
       //H1
       "DB_M256F_Scada".tAlm.tS.tS0.x0 := "M256_Manag_IDB".M256F_IDB[0].tALM.tS.x0;
       "DB_M256F_Scada".tAlm.tS.tS0.x1 := "M256_Manag_IDB".M256F_IDB[0].tALM.tS.x1;
       "DB_M256F_Scada".tAlm.tS.tS0.x2 := "M256_Manag_IDB".M256F_IDB[0].tALM.tS.x2;
       "DB_M256F_Scada".tAlm.tS.tS0.x3 := "M256_Manag_IDB".M256F_IDB[0].tALM.tS.x3;
       "DB_M256F_Scada".tAlm.tS.tS0.x4 := "M256_Manag_IDB".M256F_IDB[0].tALM.tS.x4;
       "DB_M256F_Scada".tAlm.tS.tS0.x5 := "M256_Manag_IDB".M256F_IDB[0].tALM.tS.x5;
       "DB_M256F_Scada".tAlm.tS.tS0.x6 := "M256_Manag_IDB".M256F_IDB[0].tALM.tS.x6;
       "DB_M256F_Scada".tAlm.tS.tS0.x7 := "M256_Manag_IDB".M256F_IDB[0].tALM.tS.x7;
       "DB_M256F_Scada".tAlm.tS.tS0.x8 := "M256_Manag_IDB".M256F_IDB[0].tALM.tS.x8;
       //H2
       "DB_M256F_Scada".tAlm.tS.tS0.x9 := "M256_Manag_IDB".M256F_IDB[1].tALM.tS.x0;
       "DB_M256F_Scada".tAlm.tS.tS0.x10 := "M256_Manag_IDB".M256F_IDB[1].tALM.tS.x1;
       "DB_M256F_Scada".tAlm.tS.tS0.x11 := "M256_Manag_IDB".M256F_IDB[1].tALM.tS.x2;
       "DB_M256F_Scada".tAlm.tS.tS0.x12 := "M256_Manag_IDB".M256F_IDB[1].tALM.tS.x3;
       "DB_M256F_Scada".tAlm.tS.tS0.x13 := "M256_Manag_IDB".M256F_IDB[1].tALM.tS.x4;
       "DB_M256F_Scada".tAlm.tS.tS0.x14 := "M256_Manag_IDB".M256F_IDB[1].tALM.tS.x5;
       "DB_M256F_Scada".tAlm.tS.tS0.x15 := "M256_Manag_IDB".M256F_IDB[1].tALM.tS.x6;
       "DB_M256F_Scada".tAlm.tS.tS0.x16 := "M256_Manag_IDB".M256F_IDB[1].tALM.tS.x7;
       "DB_M256F_Scada".tAlm.tS.tS0.x17 := "M256_Manag_IDB".M256F_IDB[1].tALM.tS.x8;
       //H3
       "DB_M256F_Scada".tAlm.tS.tS0.x18 := "M256_Manag_IDB".M256F_IDB[2].tALM.tS.x0;
       "DB_M256F_Scada".tAlm.tS.tS0.x19 := "M256_Manag_IDB".M256F_IDB[2].tALM.tS.x1;
       "DB_M256F_Scada".tAlm.tS.tS0.x20 := "M256_Manag_IDB".M256F_IDB[2].tALM.tS.x2;
       "DB_M256F_Scada".tAlm.tS.tS0.x21 := "M256_Manag_IDB".M256F_IDB[2].tALM.tS.x3;
       "DB_M256F_Scada".tAlm.tS.tS0.x22 := "M256_Manag_IDB".M256F_IDB[2].tALM.tS.x4;
       "DB_M256F_Scada".tAlm.tS.tS0.x23 := "M256_Manag_IDB".M256F_IDB[2].tALM.tS.x5;
       "DB_M256F_Scada".tAlm.tS.tS0.x24 := "M256_Manag_IDB".M256F_IDB[2].tALM.tS.x6;
       "DB_M256F_Scada".tAlm.tS.tS0.x25 := "M256_Manag_IDB".M256F_IDB[2].tALM.tS.x7;
       "DB_M256F_Scada".tAlm.tS.tS0.x26 := "M256_Manag_IDB".M256F_IDB[2].tALM.tS.x8;
       //H4
       "DB_M256F_Scada".tAlm.tS.tS1.x0 := "M256_Manag_IDB".M256F_IDB[3].tALM.tS.x0;
       "DB_M256F_Scada".tAlm.tS.tS1.x1 := "M256_Manag_IDB".M256F_IDB[3].tALM.tS.x1;
       "DB_M256F_Scada".tAlm.tS.tS1.x2 := "M256_Manag_IDB".M256F_IDB[3].tALM.tS.x2;
       "DB_M256F_Scada".tAlm.tS.tS1.x3 := "M256_Manag_IDB".M256F_IDB[3].tALM.tS.x3;
       "DB_M256F_Scada".tAlm.tS.tS1.x4 := "M256_Manag_IDB".M256F_IDB[3].tALM.tS.x4;
       "DB_M256F_Scada".tAlm.tS.tS1.x5 := "M256_Manag_IDB".M256F_IDB[3].tALM.tS.x5;
       "DB_M256F_Scada".tAlm.tS.tS1.x6 := "M256_Manag_IDB".M256F_IDB[3].tALM.tS.x6;
       "DB_M256F_Scada".tAlm.tS.tS1.x7 := "M256_Manag_IDB".M256F_IDB[3].tALM.tS.x7;
       "DB_M256F_Scada".tAlm.tS.tS1.x8 := "M256_Manag_IDB".M256F_IDB[3].tALM.tS.x8;
       //H5
       "DB_M256F_Scada".tAlm.tS.tS1.x9 := "M256_Manag_IDB".M256F_IDB[4].tALM.tS.x0;
       "DB_M256F_Scada".tAlm.tS.tS1.x10 := "M256_Manag_IDB".M256F_IDB[4].tALM.tS.x1;
       "DB_M256F_Scada".tAlm.tS.tS1.x11 := "M256_Manag_IDB".M256F_IDB[4].tALM.tS.x2;
       "DB_M256F_Scada".tAlm.tS.tS1.x12 := "M256_Manag_IDB".M256F_IDB[4].tALM.tS.x3;
       "DB_M256F_Scada".tAlm.tS.tS1.x13 := "M256_Manag_IDB".M256F_IDB[4].tALM.tS.x4;
       "DB_M256F_Scada".tAlm.tS.tS1.x14 := "M256_Manag_IDB".M256F_IDB[4].tALM.tS.x5;
       "DB_M256F_Scada".tAlm.tS.tS1.x15 := "M256_Manag_IDB".M256F_IDB[4].tALM.tS.x6;
       "DB_M256F_Scada".tAlm.tS.tS1.x16 := "M256_Manag_IDB".M256F_IDB[4].tALM.tS.x7;
       "DB_M256F_Scada".tAlm.tS.tS1.x17 := "M256_Manag_IDB".M256F_IDB[4].tALM.tS.x8;
       //H6
       "DB_M256F_Scada".tAlm.tS.tS1.x18 := "M256_Manag_IDB".M256F_IDB[5].tALM.tS.x0;
       "DB_M256F_Scada".tAlm.tS.tS1.x19 := "M256_Manag_IDB".M256F_IDB[5].tALM.tS.x1;
       "DB_M256F_Scada".tAlm.tS.tS1.x20 := "M256_Manag_IDB".M256F_IDB[5].tALM.tS.x2;
       "DB_M256F_Scada".tAlm.tS.tS1.x21 := "M256_Manag_IDB".M256F_IDB[5].tALM.tS.x3;
       "DB_M256F_Scada".tAlm.tS.tS1.x22 := "M256_Manag_IDB".M256F_IDB[5].tALM.tS.x4;
       "DB_M256F_Scada".tAlm.tS.tS1.x23 := "M256_Manag_IDB".M256F_IDB[5].tALM.tS.x5;
       "DB_M256F_Scada".tAlm.tS.tS1.x24 := "M256_Manag_IDB".M256F_IDB[5].tALM.tS.x6;
       "DB_M256F_Scada".tAlm.tS.tS1.x25 := "M256_Manag_IDB".M256F_IDB[5].tALM.tS.x7;
       "DB_M256F_Scada".tAlm.tS.tS1.x26 := "M256_Manag_IDB".M256F_IDB[5].tALM.tS.x8;
       //H7
       "DB_M256F_Scada".tAlm.tS.tS2.x0 := "M256_Manag_IDB".M256F_IDB[6].tALM.tS.x0;
       "DB_M256F_Scada".tAlm.tS.tS2.x1 := "M256_Manag_IDB".M256F_IDB[6].tALM.tS.x1;
       "DB_M256F_Scada".tAlm.tS.tS2.x2 := "M256_Manag_IDB".M256F_IDB[6].tALM.tS.x2;
       "DB_M256F_Scada".tAlm.tS.tS2.x3 := "M256_Manag_IDB".M256F_IDB[6].tALM.tS.x3;
       "DB_M256F_Scada".tAlm.tS.tS2.x4 := "M256_Manag_IDB".M256F_IDB[6].tALM.tS.x4;
       "DB_M256F_Scada".tAlm.tS.tS2.x5 := "M256_Manag_IDB".M256F_IDB[6].tALM.tS.x5;
       "DB_M256F_Scada".tAlm.tS.tS2.x6 := "M256_Manag_IDB".M256F_IDB[6].tALM.tS.x6;
       "DB_M256F_Scada".tAlm.tS.tS2.x7 := "M256_Manag_IDB".M256F_IDB[6].tALM.tS.x7;
       "DB_M256F_Scada".tAlm.tS.tS2.x8 := "M256_Manag_IDB".M256F_IDB[6].tALM.tS.x8;
       //H8
       "DB_M256F_Scada".tAlm.tS.tS2.x9 := "M256_Manag_IDB".M256F_IDB[7].tALM.tS.x0;
       "DB_M256F_Scada".tAlm.tS.tS2.x10 := "M256_Manag_IDB".M256F_IDB[7].tALM.tS.x1;
       "DB_M256F_Scada".tAlm.tS.tS2.x11 := "M256_Manag_IDB".M256F_IDB[7].tALM.tS.x2;
       "DB_M256F_Scada".tAlm.tS.tS2.x12 := "M256_Manag_IDB".M256F_IDB[7].tALM.tS.x3;
       "DB_M256F_Scada".tAlm.tS.tS2.x13 := "M256_Manag_IDB".M256F_IDB[7].tALM.tS.x4;
       "DB_M256F_Scada".tAlm.tS.tS2.x14 := "M256_Manag_IDB".M256F_IDB[7].tALM.tS.x5;
       "DB_M256F_Scada".tAlm.tS.tS2.x15 := "M256_Manag_IDB".M256F_IDB[7].tALM.tS.x6;
       "DB_M256F_Scada".tAlm.tS.tS2.x16 := "M256_Manag_IDB".M256F_IDB[7].tALM.tS.x7;
       "DB_M256F_Scada".tAlm.tS.tS2.x17 := "M256_Manag_IDB".M256F_IDB[7].tALM.tS.x8;



       //Move ARMING HMR
       //H1
       "DB_M256A_Scada".tHMR.dHeadStatus_H1 := "M256_Manag_IDB".M256A_IDB[0].tHMR.dHeadStatus;
       "DB_M256A_Scada".tHMR.tManCmd.xMan_DescentFdbk_H1:="M256_Manag_IDB".M256A_IDB[0].tHMR.tManCmd.xMan_DescentFdbk;
       "DB_M256A_Scada".tHMR.tManCmd.xMan_RiseFdbk_H1 := "M256_Manag_IDB".M256A_IDB[0].tHMR.tManCmd.xMan_RiseFdbk;
       //H2
       "DB_M256A_Scada".tHMR.dHeadStatus_H2 := "M256_Manag_IDB".M256A_IDB[1].tHMR.dHeadStatus;
       "DB_M256A_Scada".tHMR.tManCmd.xMan_DescentFdbk_H2 := "M256_Manag_IDB".M256A_IDB[1].tHMR.tManCmd.xMan_DescentFdbk;
       "DB_M256A_Scada".tHMR.tManCmd.xMan_RiseFdbk_H2 := "M256_Manag_IDB".M256A_IDB[1].tHMR.tManCmd.xMan_RiseFdbk;
       //H3
       "DB_M256A_Scada".tHMR.dHeadStatus_H3 := "M256_Manag_IDB".M256A_IDB[2].tHMR.dHeadStatus;
       "DB_M256A_Scada".tHMR.tManCmd.xMan_DescentFdbk_H3 := "M256_Manag_IDB".M256A_IDB[2].tHMR.tManCmd.xMan_DescentFdbk;
       "DB_M256A_Scada".tHMR.tManCmd.xMan_RiseFdbk_H3 := "M256_Manag_IDB".M256A_IDB[2].tHMR.tManCmd.xMan_RiseFdbk;
       //H4
       "DB_M256A_Scada".tHMR.dHeadStatus_H4 := "M256_Manag_IDB".M256A_IDB[3].tHMR.dHeadStatus;
       "DB_M256A_Scada".tHMR.tManCmd.xMan_DescentFdbk_H4 := "M256_Manag_IDB".M256A_IDB[3].tHMR.tManCmd.xMan_DescentFdbk;
       "DB_M256A_Scada".tHMR.tManCmd.xMan_RiseFdbk_H4 := "M256_Manag_IDB".M256A_IDB[3].tHMR.tManCmd.xMan_RiseFdbk;
       //H5
       "DB_M256A_Scada".tHMR.dHeadStatus_H5 := "M256_Manag_IDB".M256A_IDB[4].tHMR.dHeadStatus;
       "DB_M256A_Scada".tHMR.tManCmd.xMan_DescentFdbk_H5 := "M256_Manag_IDB".M256A_IDB[4].tHMR.tManCmd.xMan_DescentFdbk;
       "DB_M256A_Scada".tHMR.tManCmd.xMan_RiseFdbk_H5 := "M256_Manag_IDB".M256A_IDB[4].tHMR.tManCmd.xMan_RiseFdbk;
       //H6
       "DB_M256A_Scada".tHMR.dHeadStatus_H6 := "M256_Manag_IDB".M256A_IDB[5].tHMR.dHeadStatus;
       "DB_M256A_Scada".tHMR.tManCmd.xMan_DescentFdbk_H6 := "M256_Manag_IDB".M256A_IDB[5].tHMR.tManCmd.xMan_DescentFdbk;
       "DB_M256A_Scada".tHMR.tManCmd.xMan_RiseFdbk_H6 := "M256_Manag_IDB".M256A_IDB[5].tHMR.tManCmd.xMan_RiseFdbk;
       //H7
       "DB_M256A_Scada".tHMR.dHeadStatus_H7 := "M256_Manag_IDB".M256A_IDB[6].tHMR.dHeadStatus;
       "DB_M256A_Scada".tHMR.tManCmd.xMan_DescentFdbk_H7 := "M256_Manag_IDB".M256A_IDB[6].tHMR.tManCmd.xMan_DescentFdbk;
       "DB_M256A_Scada".tHMR.tManCmd.xMan_RiseFdbk_H7 := "M256_Manag_IDB".M256A_IDB[6].tHMR.tManCmd.xMan_RiseFdbk;
       //H8
       "DB_M256A_Scada".tHMR.dHeadStatus_H8 := "M256_Manag_IDB".M256A_IDB[7].tHMR.dHeadStatus;
       "DB_M256A_Scada".tHMR.tManCmd.xMan_DescentFdbk_H8 := "M256_Manag_IDB".M256A_IDB[7].tHMR.tManCmd.xMan_DescentFdbk;
       "DB_M256A_Scada".tHMR.tManCmd.xMan_RiseFdbk_H8 := "M256_Manag_IDB".M256A_IDB[7].tHMR.tManCmd.xMan_RiseFdbk;

       //Move ARMING HMW
       //H1
       "M256_Manag_IDB".M256A_IDB[0].tHMW.dDescentReactTime_ms:="DB_M256A_Scada".tHMW.dDescentReactTime_ms_H1;
       "M256_Manag_IDB".M256A_IDB[0].tHMW.dRaiseReactTime_ms := "DB_M256A_Scada".tHMW.dRaiseReactTime_ms_H1;
       "M256_Manag_IDB".M256A_IDB[0].tHMW.tManCmd.xManDescent := "DB_M256A_Scada".tHMW.tManCmd.xManDescent_H1;
       "M256_Manag_IDB".M256A_IDB[0].tHMW.tManCmd.xManRise := "DB_M256A_Scada".tHMW.tManCmd.xManRise_H1;
       //H2
       "M256_Manag_IDB".M256A_IDB[1].tHMW.dDescentReactTime_ms := "DB_M256A_Scada".tHMW.dDescentReactTime_ms_H2;
       "M256_Manag_IDB".M256A_IDB[1].tHMW.dRaiseReactTime_ms := "DB_M256A_Scada".tHMW.dRaiseReactTime_ms_H2;
       "M256_Manag_IDB".M256A_IDB[1].tHMW.tManCmd.xManDescent := "DB_M256A_Scada".tHMW.tManCmd.xManDescent_H2;
       "M256_Manag_IDB".M256A_IDB[1].tHMW.tManCmd.xManRise := "DB_M256A_Scada".tHMW.tManCmd.xManRise_H2;
       //H3
       "M256_Manag_IDB".M256A_IDB[2].tHMW.dDescentReactTime_ms := "DB_M256A_Scada".tHMW.dDescentReactTime_ms_H3;
       "M256_Manag_IDB".M256A_IDB[2].tHMW.dRaiseReactTime_ms := "DB_M256A_Scada".tHMW.dRaiseReactTime_ms_H3;
       "M256_Manag_IDB".M256A_IDB[2].tHMW.tManCmd.xManDescent := "DB_M256A_Scada".tHMW.tManCmd.xManDescent_H3;
       "M256_Manag_IDB".M256A_IDB[2].tHMW.tManCmd.xManRise := "DB_M256A_Scada".tHMW.tManCmd.xManRise_H3;
       //H4
       "M256_Manag_IDB".M256A_IDB[3].tHMW.dDescentReactTime_ms := "DB_M256A_Scada".tHMW.dDescentReactTime_ms_H4;
       "M256_Manag_IDB".M256A_IDB[3].tHMW.dRaiseReactTime_ms := "DB_M256A_Scada".tHMW.dRaiseReactTime_ms_H4;
       "M256_Manag_IDB".M256A_IDB[3].tHMW.tManCmd.xManDescent := "DB_M256A_Scada".tHMW.tManCmd.xManDescent_H4;
       "M256_Manag_IDB".M256A_IDB[3].tHMW.tManCmd.xManRise := "DB_M256A_Scada".tHMW.tManCmd.xManRise_H4;
       //H5
       "M256_Manag_IDB".M256A_IDB[4].tHMW.dDescentReactTime_ms := "DB_M256A_Scada".tHMW.dDescentReactTime_ms_H5;
       "M256_Manag_IDB".M256A_IDB[4].tHMW.dRaiseReactTime_ms := "DB_M256A_Scada".tHMW.dRaiseReactTime_ms_H5;
       "M256_Manag_IDB".M256A_IDB[4].tHMW.tManCmd.xManDescent := "DB_M256A_Scada".tHMW.tManCmd.xManDescent_H5;
       "M256_Manag_IDB".M256A_IDB[4].tHMW.tManCmd.xManRise := "DB_M256A_Scada".tHMW.tManCmd.xManRise_H5;
       //H6
       "M256_Manag_IDB".M256A_IDB[5].tHMW.dDescentReactTime_ms := "DB_M256A_Scada".tHMW.dDescentReactTime_ms_H6;
       "M256_Manag_IDB".M256A_IDB[5].tHMW.dRaiseReactTime_ms := "DB_M256A_Scada".tHMW.dRaiseReactTime_ms_H6;
       "M256_Manag_IDB".M256A_IDB[5].tHMW.tManCmd.xManDescent := "DB_M256A_Scada".tHMW.tManCmd.xManDescent_H6;
       "M256_Manag_IDB".M256A_IDB[5].tHMW.tManCmd.xManRise := "DB_M256A_Scada".tHMW.tManCmd.xManRise_H6;
       //H7
       "M256_Manag_IDB".M256A_IDB[6].tHMW.dDescentReactTime_ms := "DB_M256A_Scada".tHMW.dDescentReactTime_ms_H7;
       "M256_Manag_IDB".M256A_IDB[6].tHMW.dRaiseReactTime_ms := "DB_M256A_Scada".tHMW.dRaiseReactTime_ms_H7;
       "M256_Manag_IDB".M256A_IDB[6].tHMW.tManCmd.xManDescent := "DB_M256A_Scada".tHMW.tManCmd.xManDescent_H7;
       "M256_Manag_IDB".M256A_IDB[6].tHMW.tManCmd.xManRise := "DB_M256A_Scada".tHMW.tManCmd.xManRise_H7;
       //H8
       "M256_Manag_IDB".M256A_IDB[7].tHMW.dDescentReactTime_ms := "DB_M256A_Scada".tHMW.dDescentReactTime_ms_H8;
       "M256_Manag_IDB".M256A_IDB[7].tHMW.dRaiseReactTime_ms := "DB_M256A_Scada".tHMW.dRaiseReactTime_ms_H8;
       "M256_Manag_IDB".M256A_IDB[7].tHMW.tManCmd.xManDescent := "DB_M256A_Scada".tHMW.tManCmd.xManDescent_H8;
       "M256_Manag_IDB".M256A_IDB[7].tHMW.tManCmd.xManRise := "DB_M256A_Scada".tHMW.tManCmd.xManRise_H8;


       //Move ARMING ALM

       "DB_M256A_Scada".tAlm.tF := "M256_Manag_IDB".M256A_IDB[0].tALM.tF;

       "DB_M256A_Scada".tAlm.tW := "M256_Manag_IDB".M256A_IDB[0].tALM.tW;

               //H1
       "DB_M256A_Scada".tAlm.tS.tS0.x0 := "M256_Manag_IDB".M256A_IDB[0].tALM.tS.xNotWorkPos;
       "DB_M256A_Scada".tAlm.tS.tS0.x1 := "M256_Manag_IDB".M256A_IDB[0].tALM.tS.x1;
       "DB_M256A_Scada".tAlm.tS.tS0.x2 := "M256_Manag_IDB".M256A_IDB[0].tALM.tS.x2;
       "DB_M256A_Scada".tAlm.tS.tS0.x3 := "M256_Manag_IDB".M256A_IDB[0].tALM.tS.x3;
       "DB_M256A_Scada".tAlm.tS.tS0.x4 := "M256_Manag_IDB".M256A_IDB[0].tALM.tS.x4;
       "DB_M256A_Scada".tAlm.tS.tS0.x5 := "M256_Manag_IDB".M256A_IDB[0].tALM.tS.x5;
       "DB_M256A_Scada".tAlm.tS.tS0.x6 := "M256_Manag_IDB".M256A_IDB[0].tALM.tS.x6;
       "DB_M256A_Scada".tAlm.tS.tS0.x7 := "M256_Manag_IDB".M256A_IDB[0].tALM.tS.x7;
       "DB_M256A_Scada".tAlm.tS.tS0.x8 := "M256_Manag_IDB".M256A_IDB[0].tALM.tS.x8;
               //H2
       "DB_M256A_Scada".tAlm.tS.tS0.x9 := "M256_Manag_IDB".M256A_IDB[1].tALM.tS.xNotWorkPos;
       "DB_M256A_Scada".tAlm.tS.tS0.x10 := "M256_Manag_IDB".M256A_IDB[1].tALM.tS.x1;
       "DB_M256A_Scada".tAlm.tS.tS0.x11 := "M256_Manag_IDB".M256A_IDB[1].tALM.tS.x2;
       "DB_M256A_Scada".tAlm.tS.tS0.x12 := "M256_Manag_IDB".M256A_IDB[1].tALM.tS.x3;
       "DB_M256A_Scada".tAlm.tS.tS0.x13 := "M256_Manag_IDB".M256A_IDB[1].tALM.tS.x4;
       "DB_M256A_Scada".tAlm.tS.tS0.x14 := "M256_Manag_IDB".M256A_IDB[1].tALM.tS.x5;
       "DB_M256A_Scada".tAlm.tS.tS0.x15 := "M256_Manag_IDB".M256A_IDB[1].tALM.tS.x6;
       "DB_M256A_Scada".tAlm.tS.tS0.x16 := "M256_Manag_IDB".M256A_IDB[1].tALM.tS.x7;
       "DB_M256A_Scada".tAlm.tS.tS0.x17 := "M256_Manag_IDB".M256A_IDB[1].tALM.tS.x8;
               //H3
       "DB_M256A_Scada".tAlm.tS.tS0.x18 := "M256_Manag_IDB".M256A_IDB[2].tALM.tS.xNotWorkPos;
       "DB_M256A_Scada".tAlm.tS.tS0.x19 := "M256_Manag_IDB".M256A_IDB[2].tALM.tS.x1;
       "DB_M256A_Scada".tAlm.tS.tS0.x20 := "M256_Manag_IDB".M256A_IDB[2].tALM.tS.x2;
       "DB_M256A_Scada".tAlm.tS.tS0.x21 := "M256_Manag_IDB".M256A_IDB[2].tALM.tS.x3;
       "DB_M256A_Scada".tAlm.tS.tS0.x22 := "M256_Manag_IDB".M256A_IDB[2].tALM.tS.x4;
       "DB_M256A_Scada".tAlm.tS.tS0.x23 := "M256_Manag_IDB".M256A_IDB[2].tALM.tS.x5;
       "DB_M256A_Scada".tAlm.tS.tS0.x24 := "M256_Manag_IDB".M256A_IDB[2].tALM.tS.x6;
       "DB_M256A_Scada".tAlm.tS.tS0.x25 := "M256_Manag_IDB".M256A_IDB[2].tALM.tS.x7;
       "DB_M256A_Scada".tAlm.tS.tS0.x26 := "M256_Manag_IDB".M256A_IDB[2].tALM.tS.x8;
               //H4
       "DB_M256A_Scada".tAlm.tS.tS1.x0 := "M256_Manag_IDB".M256A_IDB[3].tALM.tS.xNotWorkPos;
       "DB_M256A_Scada".tAlm.tS.tS1.x1 := "M256_Manag_IDB".M256A_IDB[3].tALM.tS.x1;
       "DB_M256A_Scada".tAlm.tS.tS1.x2 := "M256_Manag_IDB".M256A_IDB[3].tALM.tS.x2;
       "DB_M256A_Scada".tAlm.tS.tS1.x3 := "M256_Manag_IDB".M256A_IDB[3].tALM.tS.x3;
       "DB_M256A_Scada".tAlm.tS.tS1.x4 := "M256_Manag_IDB".M256A_IDB[3].tALM.tS.x4;
       "DB_M256A_Scada".tAlm.tS.tS1.x5 := "M256_Manag_IDB".M256A_IDB[3].tALM.tS.x5;
       "DB_M256A_Scada".tAlm.tS.tS1.x6 := "M256_Manag_IDB".M256A_IDB[3].tALM.tS.x6;
       "DB_M256A_Scada".tAlm.tS.tS1.x7 := "M256_Manag_IDB".M256A_IDB[3].tALM.tS.x7;
       "DB_M256A_Scada".tAlm.tS.tS1.x8 := "M256_Manag_IDB".M256A_IDB[3].tALM.tS.x8;
               //H5
       "DB_M256A_Scada".tAlm.tS.tS1.x9 := "M256_Manag_IDB".M256A_IDB[4].tALM.tS.xNotWorkPos;
       "DB_M256A_Scada".tAlm.tS.tS1.x10 := "M256_Manag_IDB".M256A_IDB[4].tALM.tS.x1;
       "DB_M256A_Scada".tAlm.tS.tS1.x11 := "M256_Manag_IDB".M256A_IDB[4].tALM.tS.x2;
       "DB_M256A_Scada".tAlm.tS.tS1.x12 := "M256_Manag_IDB".M256A_IDB[4].tALM.tS.x3;
       "DB_M256A_Scada".tAlm.tS.tS1.x13 := "M256_Manag_IDB".M256A_IDB[4].tALM.tS.x4;
       "DB_M256A_Scada".tAlm.tS.tS1.x14 := "M256_Manag_IDB".M256A_IDB[4].tALM.tS.x5;
       "DB_M256A_Scada".tAlm.tS.tS1.x15 := "M256_Manag_IDB".M256A_IDB[4].tALM.tS.x6;
       "DB_M256A_Scada".tAlm.tS.tS1.x16 := "M256_Manag_IDB".M256A_IDB[4].tALM.tS.x7;
       "DB_M256A_Scada".tAlm.tS.tS1.x17 := "M256_Manag_IDB".M256A_IDB[4].tALM.tS.x8;
               //H6
       "DB_M256A_Scada".tAlm.tS.tS1.x18 := "M256_Manag_IDB".M256A_IDB[5].tALM.tS.xNotWorkPos;
       "DB_M256A_Scada".tAlm.tS.tS1.x19 := "M256_Manag_IDB".M256A_IDB[5].tALM.tS.x1;
       "DB_M256A_Scada".tAlm.tS.tS1.x20 := "M256_Manag_IDB".M256A_IDB[5].tALM.tS.x2;
       "DB_M256A_Scada".tAlm.tS.tS1.x21 := "M256_Manag_IDB".M256A_IDB[5].tALM.tS.x3;
       "DB_M256A_Scada".tAlm.tS.tS1.x22 := "M256_Manag_IDB".M256A_IDB[5].tALM.tS.x4;
       "DB_M256A_Scada".tAlm.tS.tS1.x23 := "M256_Manag_IDB".M256A_IDB[5].tALM.tS.x5;
       "DB_M256A_Scada".tAlm.tS.tS1.x24 := "M256_Manag_IDB".M256A_IDB[5].tALM.tS.x6;
       "DB_M256A_Scada".tAlm.tS.tS1.x25 := "M256_Manag_IDB".M256A_IDB[5].tALM.tS.x7;
       "DB_M256A_Scada".tAlm.tS.tS1.x26 := "M256_Manag_IDB".M256A_IDB[5].tALM.tS.x8;
               //H7
       "DB_M256A_Scada".tAlm.tS.tS2.x0 := "M256_Manag_IDB".M256A_IDB[6].tALM.tS.xNotWorkPos;
       "DB_M256A_Scada".tAlm.tS.tS2.x1 := "M256_Manag_IDB".M256A_IDB[6].tALM.tS.x1;
       "DB_M256A_Scada".tAlm.tS.tS2.x2 := "M256_Manag_IDB".M256A_IDB[6].tALM.tS.x2;
       "DB_M256A_Scada".tAlm.tS.tS2.x3 := "M256_Manag_IDB".M256A_IDB[6].tALM.tS.x3;
       "DB_M256A_Scada".tAlm.tS.tS2.x4 := "M256_Manag_IDB".M256A_IDB[6].tALM.tS.x4;
       "DB_M256A_Scada".tAlm.tS.tS2.x5 := "M256_Manag_IDB".M256A_IDB[6].tALM.tS.x5;
       "DB_M256A_Scada".tAlm.tS.tS2.x6 := "M256_Manag_IDB".M256A_IDB[6].tALM.tS.x6;
       "DB_M256A_Scada".tAlm.tS.tS2.x7 := "M256_Manag_IDB".M256A_IDB[6].tALM.tS.x7;
       "DB_M256A_Scada".tAlm.tS.tS2.x8 := "M256_Manag_IDB".M256A_IDB[6].tALM.tS.x8;
               //H8
       "DB_M256A_Scada".tAlm.tS.tS2.x9 := "M256_Manag_IDB".M256A_IDB[7].tALM.tS.xNotWorkPos;
       "DB_M256A_Scada".tAlm.tS.tS2.x10 := "M256_Manag_IDB".M256A_IDB[7].tALM.tS.x1;
       "DB_M256A_Scada".tAlm.tS.tS2.x11 := "M256_Manag_IDB".M256A_IDB[7].tALM.tS.x2;
       "DB_M256A_Scada".tAlm.tS.tS2.x12 := "M256_Manag_IDB".M256A_IDB[7].tALM.tS.x3;
       "DB_M256A_Scada".tAlm.tS.tS2.x13 := "M256_Manag_IDB".M256A_IDB[7].tALM.tS.x4;
       "DB_M256A_Scada".tAlm.tS.tS2.x14 := "M256_Manag_IDB".M256A_IDB[7].tALM.tS.x5;
       "DB_M256A_Scada".tAlm.tS.tS2.x15 := "M256_Manag_IDB".M256A_IDB[7].tALM.tS.x6;
       "DB_M256A_Scada".tAlm.tS.tS2.x16 := "M256_Manag_IDB".M256A_IDB[7].tALM.tS.x7;
       "DB_M256A_Scada".tAlm.tS.tS2.x17 := "M256_Manag_IDB".M256A_IDB[7].tALM.tS.x8;
END_FUNCTION

// folder: Communication

FUNCTION "CM_Management" : Void   // FC14, LAD
{ S7_Optimized_Access := 'TRUE' }
VERSION : 0.1
   VAR_TEMP
      TMP_dDummy : DInt;
   END_VAR
   VAR_TEMP   // added for the SCL form of the ladder/FBD networks
      _w1 : Bool;
   END_VAR
BEGIN

REGION Network 1: COSTANTS
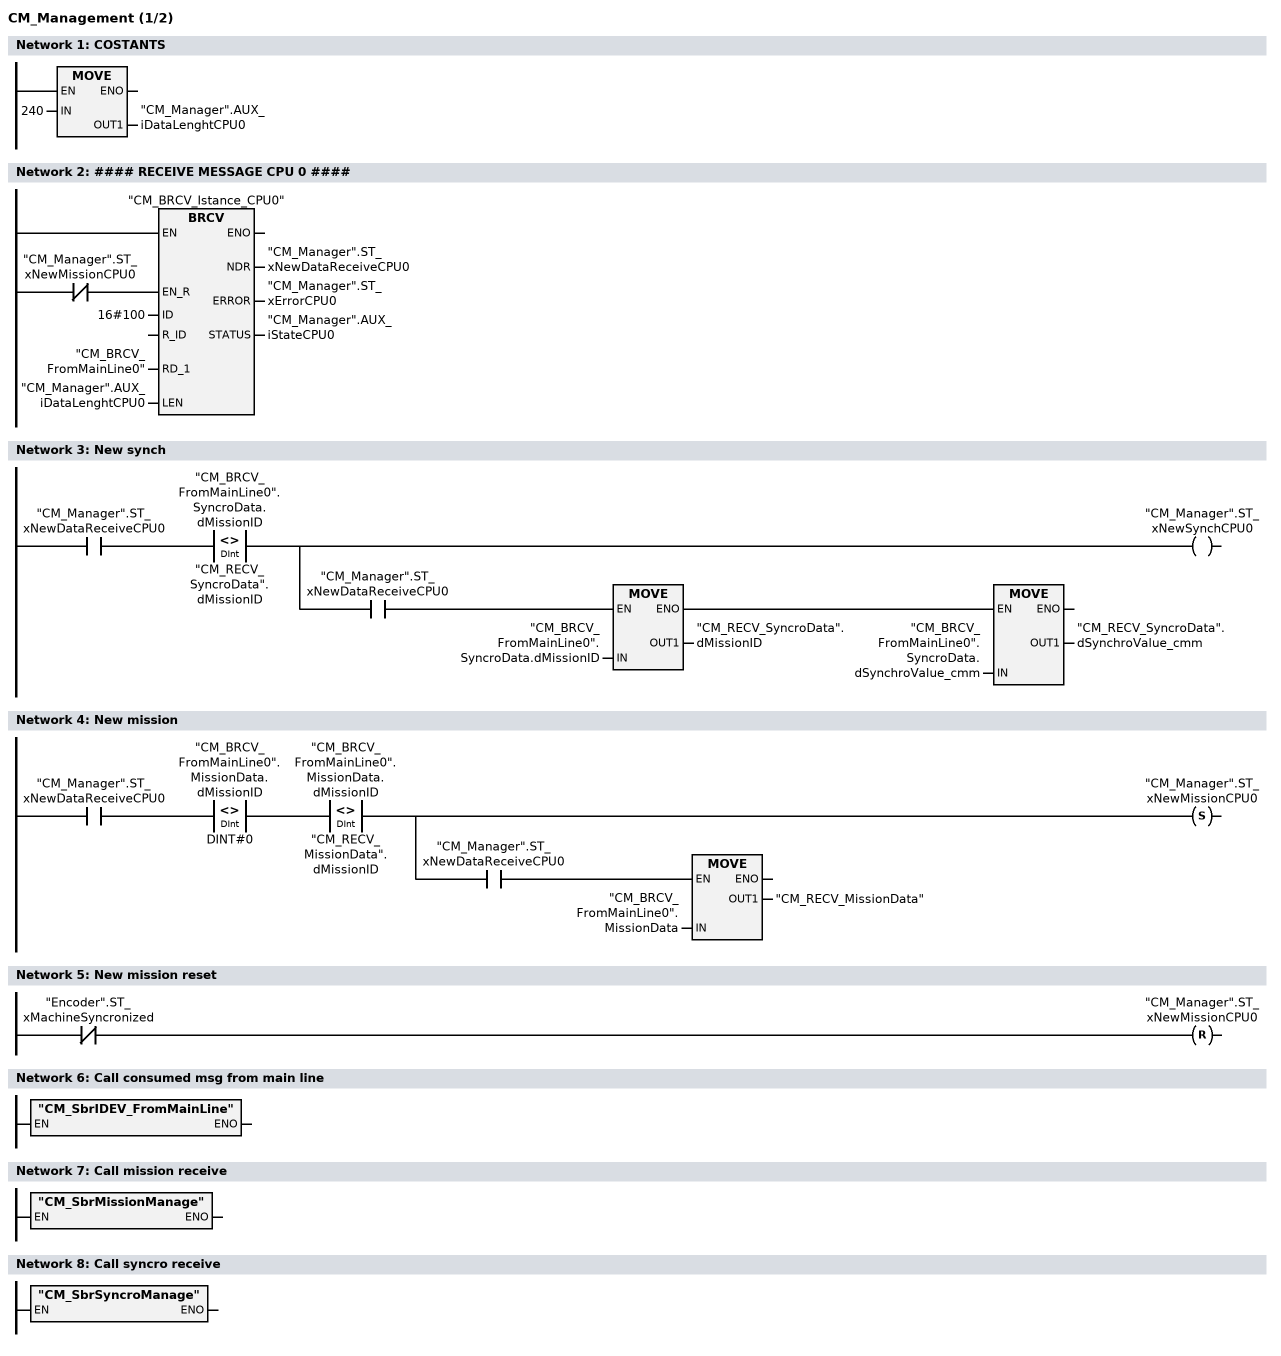
   RUNG wire#powerrail
      Move(in := 240, out1 => "CM_Manager".AUX_iDataLenghtCPU0)
   END_RUNG
   // the same network as SCL:
   "CM_Manager".AUX_iDataLenghtCPU0 := 240;
END_REGION

REGION Network 2: #### RECEIVE MESSAGE CPU 0 ####
   "CM_BRCV_Istance_CPU0"(EN_R := NOT "CM_Manager".ST_xNewMissionCPU0,   // BRCV
                          ID := 16#100,
                          RD_1 := "CM_BRCV_FromMainLine0",
                          LEN := "CM_Manager".AUX_iDataLenghtCPU0,
                          NDR => "CM_Manager".ST_xNewDataReceiveCPU0,
                          ERROR => "CM_Manager".ST_xErrorCPU0,
                          STATUS => "CM_Manager".AUX_iStateCPU0);
END_REGION

REGION Network 3: New synch
   RUNG wire#powerrail
      Contact( "CM_Manager".ST_xNewDataReceiveCPU0 )
      { S7_Templates := "SrcType := DInt" } NE_Contact(in1 := "CM_BRCV_FromMainLine0".SyncroData.dMissionID, in2 := "CM_RECV_SyncroData".dMissionID)
      wire#w1
      Coil( "CM_Manager".ST_xNewSynchCPU0 )
   END_RUNG
   RUNG wire#w1
      Contact( "CM_Manager".ST_xNewDataReceiveCPU0 )
      Move(in := "CM_BRCV_FromMainLine0".SyncroData.dMissionID, out1 => "CM_RECV_SyncroData".dMissionID)
      Move(in := "CM_BRCV_FromMainLine0".SyncroData.dSynchroValue_cmm, out1 => "CM_RECV_SyncroData".dSynchroValue_cmm)
   END_RUNG
   // the same network as SCL:
   "CM_Manager".ST_xNewSynchCPU0 := "CM_Manager".ST_xNewDataReceiveCPU0 AND ("CM_BRCV_FromMainLine0".SyncroData.dMissionID <> "CM_RECV_SyncroData".dMissionID);
   IF "CM_Manager".ST_xNewSynchCPU0 AND "CM_Manager".ST_xNewDataReceiveCPU0 THEN
       "CM_RECV_SyncroData".dMissionID := "CM_BRCV_FromMainLine0".SyncroData.dMissionID;
       "CM_RECV_SyncroData".dSynchroValue_cmm := "CM_BRCV_FromMainLine0".SyncroData.dSynchroValue_cmm;
   END_IF;
END_REGION

REGION Network 4: New mission
   RUNG wire#powerrail
      Contact( "CM_Manager".ST_xNewDataReceiveCPU0 )
      { S7_Templates := "SrcType := DInt" } NE_Contact(in1 := "CM_BRCV_FromMainLine0".MissionData.dMissionID, in2 := DINT#0)
      { S7_Templates := "SrcType := DInt" } NE_Contact(in1 := "CM_BRCV_FromMainLine0".MissionData.dMissionID, in2 := "CM_RECV_MissionData".dMissionID)
      wire#w1
      S_Coil( "CM_Manager".ST_xNewMissionCPU0 )
   END_RUNG
   RUNG wire#w1
      Contact( "CM_Manager".ST_xNewDataReceiveCPU0 )
      Move(in := "CM_BRCV_FromMainLine0".MissionData, out1 => "CM_RECV_MissionData")
   END_RUNG
   // the same network as SCL:
   #_w1 := "CM_Manager".ST_xNewDataReceiveCPU0 AND ("CM_BRCV_FromMainLine0".MissionData.dMissionID <> DINT#0) AND ("CM_BRCV_FromMainLine0".MissionData.dMissionID <> "CM_RECV_MissionData".dMissionID);
   IF #_w1 THEN "CM_Manager".ST_xNewMissionCPU0 := TRUE; END_IF;
   IF #_w1 AND "CM_Manager".ST_xNewDataReceiveCPU0 THEN
       "CM_RECV_MissionData" := "CM_BRCV_FromMainLine0".MissionData;
   END_IF;
END_REGION

REGION Network 5: New mission reset
   RUNG wire#powerrail
      I_Contact( "Encoder".ST_xMachineSyncronized )
      R_Coil( "CM_Manager".ST_xNewMissionCPU0 )
   END_RUNG
   // the same network as SCL:
   IF NOT "Encoder".ST_xMachineSyncronized THEN "CM_Manager".ST_xNewMissionCPU0 := FALSE; END_IF;
END_REGION

REGION Network 6: Call consumed msg from main line
   RUNG wire#powerrail
      "CM_SbrIDEV_FromMainLine"()
   END_RUNG
   // the same network as SCL:
   "CM_SbrIDEV_FromMainLine"();
END_REGION

REGION Network 7: Call mission receive
   RUNG wire#powerrail
      "CM_SbrMissionManage"()
   END_RUNG
   // the same network as SCL:
   "CM_SbrMissionManage"();
END_REGION

REGION Network 8: Call syncro receive
   RUNG wire#powerrail
      "CM_SbrSyncroManage"()
   END_RUNG
   // the same network as SCL:
   "CM_SbrSyncroManage"();
END_REGION

REGION Network 9: Call produced message to main line
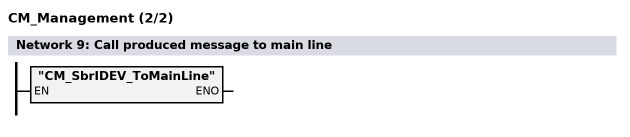
   RUNG wire#powerrail
      "CM_SbrIDEV_ToMainLine"()
   END_RUNG
   // the same network as SCL:
   "CM_SbrIDEV_ToMainLine"();
END_REGION
END_FUNCTION

FUNCTION "CM_SbrIDEV_FromMainLine" : Void   // FC15, SCL
{ S7_Optimized_Access := 'TRUE' }
VERSION : 0.1
BEGIN
   ////--------------------------------------------------------------------------------------------------------------------
   //   Copyright (c)  Bottero Spa
   //--------------------------------------------------------------
   //   Routine: ConsumedMainLine
   //       Author: Alberto Cigliutti
   //   Created: July 2016
   //--------------------------------------------------------------
   //   Description: Main line consumed message 
   //
   //   History:
   //
   ////--------------------------------------------------------------------------------------------------------------------


           "Z256".ST_xGlassBreak := "CM_IDEV_FromMainLine".xGlassBreak;
           "Z256".ST_xCycleON := "CM_IDEV_FromMainLine".xCycleON;

           IF "CM_IDEV_FromMainLine".xResetBuffers THEN
               "Z256_Manager".tInputData.xSystemReset := 1;
               "Encoder".ST_xSystemReset := 1;
           END_IF;

           IF "CM_IDEV_FromMainLine".xResetAnomaly THEN
               "Z256_hmi".tHMW.xFaultsReset := 1;
           END_IF;

    //   END_IF;
END_FUNCTION

FUNCTION "CM_SbrMissionManage" : Void   // FC16, SCL
{ S7_Optimized_Access := 'TRUE' }
VERSION : 0.1
   VAR_TEMP
      TMP_dIndex : DInt;
   END_VAR
BEGIN
   ////--------------------------------------------------------------------------------------------------------------------
   //   Copyright (c)  Bottero Spa
   //--------------------------------------------------------------
   //   Routine: CM_MissionManage
   //       Author: Alberto Cigliutti
   //   Created: July 2016
   //--------------------------------------------------------------
   //   Description: Manage the receive message
   //
   //   History:
   //
   ////--------------------------------------------------------------------------------------------------------------------

   //PLC A

   IF "CM_Manager".ST_xNewMissionCPU0 AND
       (NOT "Z256_Manager".tInputData.xNewMission) THEN


       IF (*("CM_RECV_MissionData".xPLCActive) AND*) ("Encoder".ST_xMachineSyncronized) THEN

           "Z256_Manager".tInputData.dMissionCode := "CM_RECV_MissionData".dMissionID;
           "Z256_Manager".tInputData.dMissionStart_cmm := "CM_RECV_MissionData".dMissionStart_cmm - "Encoder".AUX_dSyncroGapMainLine_cmm;
           "Z256_Manager".tInputData.dMissionEnd_cmm := "CM_RECV_MissionData".dMissionEnd_cmm - "Encoder".AUX_dSyncroGapMainLine_cmm;

           FOR #TMP_dIndex:=0 TO "CONST_dNumberOfHeadsCycle" DO
               "Z256_Manager".tInputData.rgxFireRequest[#TMP_dIndex] := "CM_RECV_MissionData".rgxFireRequest[#TMP_dIndex];
               "Z256_Manager".tInputData.rgdHeadsPosition_cmm[#TMP_dIndex] := "CM_RECV_MissionData".rgdHeadsPosition_cmm[#TMP_dIndex];
           END_FOR;

           "Z256_Manager".tInputData.xNewMission := 1;
       END_IF;

   END_IF;
END_FUNCTION

FUNCTION "CM_SbrIDEV_ToMainLine" : Void   // FC17, SCL
{ S7_Optimized_Access := 'TRUE' }
VERSION : 0.1
   VAR_TEMP
      TMP_dIndex : DInt;
   END_VAR
BEGIN
   ////--------------------------------------------------------------------------------------------------------------------
   //   Copyright (c)  Bottero Spa
   //--------------------------------------------------------------
   //   Routine: ProducedMainLine          
   //       Author: Alberto Cigliutti
   //   Created: July 2016
   //--------------------------------------------------------------
   //   Description:
   //
   //   History:
   //
   ////--------------------------------------------------------------------------------------------------------------------

   //Send request information to main line

   //Glass break in progress
   "CM_IDEV_ToMainLine".rgxStatus[0] := "CM_IDEV_FromMainLine".xGlassBreak AND (NOT "Z256_hmi".tHMW.xCutOnBreakEnabled);

   //Heads up button engaged
   "CM_IDEV_ToMainLine".rgxStatus[1] := "M256_Manag_IDB".M256A_IDB[0].INPUT_xHeadsUpIstan;

   //Bridge enabled
   "CM_IDEV_ToMainLine".rgxStatus[2] := TRUE;
   IF "M256_Manag_IDB".M256A_ST_xAllHeadStoppingFaults OR "M256_Manag_IDB".M256F_ST_xAllHeadStoppingFaults OR "M256_Manag_IDB".M256M_ST_xAllHeadStoppingFaults
       (*OR "Z256_HMI".tHMR.dProdModeActual<>3*) THEN
       "CM_IDEV_ToMainLine".rgxStatus[2] := FALSE;
   END_IF;

   //Bridge locked
   "CM_IDEV_ToMainLine".rgxStatus[3] := FALSE;

   //Cut offset calibration request (NOT USED ON MAIN LINE)
   "CM_IDEV_ToMainLine".rgxStatus[8] := FALSE;

   FOR #TMP_dIndex := 0 TO "CONST_dNumberOfHeadsCycle" DO
       "CM_IDEV_ToMainLine".rgdHeadsPositions_cmm[#TMP_dIndex] := "M256_Manag_IDB".M256M_IDB[#TMP_dIndex].AUX_dHeadActualPosition_cmm;
       "CM_IDEV_ToMainLine".rgxHeadStatus[#TMP_dIndex] := "M256_Manag_IDB".M256M_ST_xAllHeadReferred AND "Z256".INPUT_rgxHeadsInProduction[#TMP_dIndex]
       AND "Z256_hmi".tHMR.dProdModeActual=3;
       "CM_IDEV_ToMainLine".rgdHeadsPressure[#TMP_dIndex] := "M256_Manag_IDB".M256F_IDB[#TMP_dIndex].tHMW.dHeadPressure_mN;
       "CM_IDEV_ToMainLine".rgrHeadsSpace[#TMP_dIndex] := "M256_Manag_IDB".M256F_IDB[#TMP_dIndex].tHMR.rHeadUsage_km;

   END_FOR;

   //stop firing OB to have consistent data
   "CM_Manager".ST_MutingFiringOB := 1;
   FOR #TMP_dIndex := 0 TO "CONST_dNumberOfHeadsCycle" DO
       "CM_Manager".AUX_rgdHeadMissionIDInProg_Copy[#TMP_dIndex] := "M256_Manag_IDB".M256F_IDB[#TMP_dIndex].AUX_dHeadMissionIDinProg;
       "CM_Manager".AUX_rgxHeadFiringMissionInProg_Copy[#TMP_dIndex] := "M256_Manag_IDB".M256F_IDB[#TMP_dIndex].AUX_xHeadFiringMissionInProgress;
   END_FOR;
   "CM_Manager".ST_MutingFiringOB := 0;

   FOR #TMP_dIndex := 0 TO "CONST_dNumberOfHeadsCycle" DO
       "CM_IDEV_ToMainLine".dProcessingIDPlate := "CM_Manager".AUX_rgdHeadMissionIDInProg_Copy[0];
       "CM_IDEV_ToMainLine".rgxCuttingStatus[#TMP_dIndex] := "M256_Manag_IDB".M256F_IDB[#TMP_dIndex].OUTPUT_xFireON;
   END_FOR;

   //All head fire offset (NOT USED ON MAIN LINE)
   "CM_IDEV_ToMainLine".iFireOffset_OFF := 0;
   "CM_IDEV_ToMainLine".iFireOffset_ON := 0;
END_FUNCTION

FUNCTION "CM_SbrSyncroManage" : Void   // FC19, SCL
{ S7_Optimized_Access := 'TRUE' }
VERSION : 0.1
BEGIN
   ////--------------------------------------------------------------------------------------------------------------------
   //   Copyright (c)  Bottero Spa
   //--------------------------------------------------------------
   //   Routine: Syncro Manage
   //       Author: Alberto Cigliutti
   //   Created: July 2016
   //--------------------------------------------------------------
   //   Description:
   //
   //   History:
   //
   ////--------------------------------------------------------------------------------------------------------------------
   //COPY THE DATA

   //Check data received from PLC A
   IF "CM_Manager".ST_xNewSynchCPU0
       AND (NOT "Encoder".AUX_xNewSyncroReceived) THEN

       //Data valid, if PLC is active read the value 
    //   IF "CM_RECV_SyncroData".xPLCActive THEN

           "Encoder".AUX_dNewSyncroValue_cmm := "CM_RECV_SyncroData".dSynchroValue_cmm;
           "Encoder".AUX_xNewSyncroReceived := 1;

    //   END_IF;

   END_IF;
END_FUNCTION

// folder: ILx2_Blocks

FUNCTION_BLOCK "ILx2T_Control"   // FB1, SCL
{ S7_Optimized_Access := 'TRUE' }